REGION Network 178: %DB59.DBW2
   RUNG wire#powerrail
      I_Contact( "Rec_Todas" )
      I_Contact( "ResumAla_Grave" )
      { S7_GenerateENO := "TRUE" } Move(in := 0, out1 => %DB59.DBW2)
   END_RUNG
   // the same network as SCL:
   IF NOT "Rec_Todas" AND NOT "ResumAla_Grave" THEN %DB59.DBW2 := 0; END_IF;
END_REGION

REGION Network 179: %DB59.DBD4
   RUNG wire#powerrail
      Contact( "Rec_Todas" )
      wire#w1
      { S7_GenerateENO := "TRUE" } Move(in := DW#16#FFFFFFFF, out1 => %DB59.DBD4)
   END_RUNG
   RUNG wire#powerrail
      Contact( "ResumAla_Grave" )
   END_RUNG wire#w1
   // the same network as SCL:
   IF "Rec_Todas" OR "ResumAla_Grave" THEN %DB59.DBD4 := DW#16#FFFFFFFF; END_IF;
END_REGION

REGION Network 180: %DB59.DBD4
   RUNG wire#powerrail
      I_Contact( "Rec_Todas" )
      I_Contact( "ResumAla_Grave" )
      { S7_GenerateENO := "TRUE" } Move(in := 0, out1 => %DB59.DBD4)
   END_RUNG
   // the same network as SCL:
   IF NOT "Rec_Todas" AND NOT "ResumAla_Grave" THEN %DB59.DBD4 := 0; END_IF;
END_REGION

REGION Network 181: %DB59.DBD8
   RUNG wire#powerrail
      Contact( "Rec_Todas" )
      wire#w1
      { S7_GenerateENO := "TRUE" } Move(in := DW#16#FFFFFFFF, out1 => %DB59.DBD8)
   END_RUNG
   RUNG wire#powerrail
      Contact( "ResumAla_Grave" )
   END_RUNG wire#w1
   // the same network as SCL:
   IF "Rec_Todas" OR "ResumAla_Grave" THEN %DB59.DBD8 := DW#16#FFFFFFFF; END_IF;
END_REGION

REGION Network 182: %DB59.DBD8
   RUNG wire#powerrail
      I_Contact( "Rec_Todas" )
      I_Contact( "ResumAla_Grave" )
      { S7_GenerateENO := "TRUE" } Move(in := 0, out1 => %DB59.DBD8)
   END_RUNG
   // the same network as SCL:
   IF NOT "Rec_Todas" AND NOT "ResumAla_Grave" THEN %DB59.DBD8 := 0; END_IF;
END_REGION

REGION Network 183: %DB59.DBD12
   RUNG wire#powerrail
      Contact( "Rec_Todas" )
      wire#w1
      { S7_GenerateENO := "TRUE" } Move(in := DW#16#FFFFFFFF, out1 => %DB59.DBD12)
   END_RUNG
   RUNG wire#powerrail
      Contact( "ResumAla_Grave" )
   END_RUNG wire#w1
   // the same network as SCL:
   IF "Rec_Todas" OR "ResumAla_Grave" THEN %DB59.DBD12 := DW#16#FFFFFFFF; END_IF;
END_REGION

REGION Network 184: %DB59.DBD12
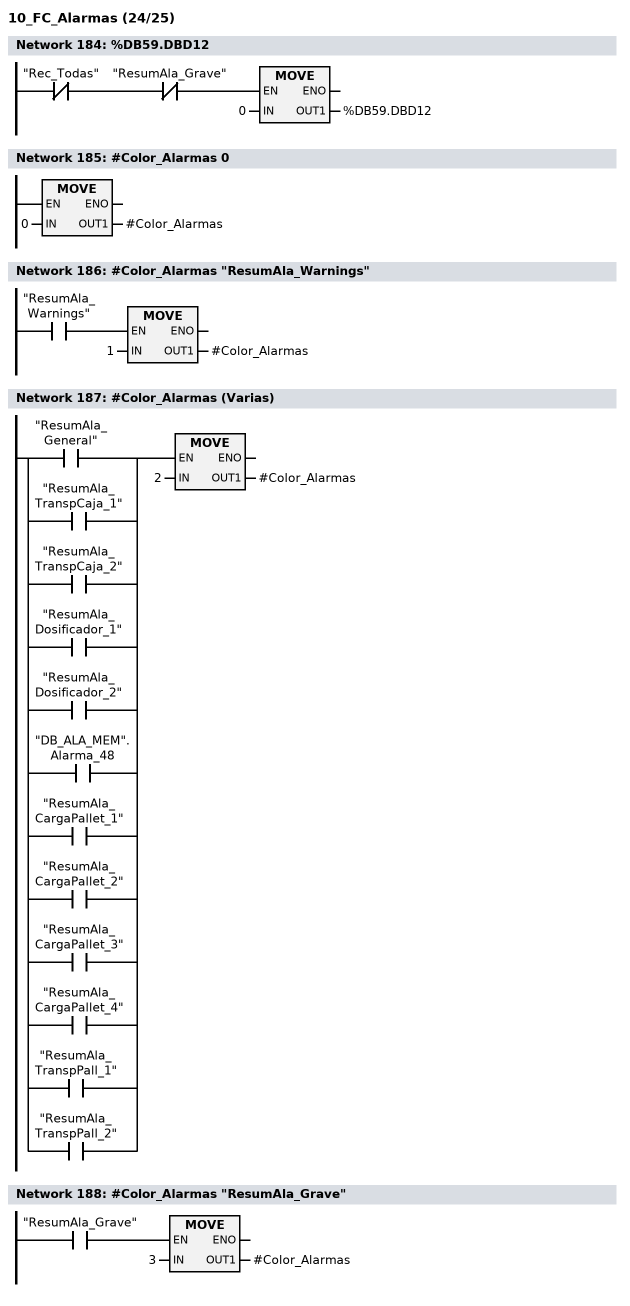
   RUNG wire#powerrail
      I_Contact( "Rec_Todas" )
      I_Contact( "ResumAla_Grave" )
      { S7_GenerateENO := "TRUE" } Move(in := 0, out1 => %DB59.DBD12)
   END_RUNG
   // the same network as SCL:
   IF NOT "Rec_Todas" AND NOT "ResumAla_Grave" THEN %DB59.DBD12 := 0; END_IF;
END_REGION

REGION Network 185: #Color_Alarmas 0
   RUNG wire#powerrail
      { S7_GenerateENO := "TRUE" } Move(in := 0, out1 => #Color_Alarmas)
   END_RUNG
   // the same network as SCL:
   #Color_Alarmas := 0;
END_REGION

REGION Network 186: #Color_Alarmas "ResumAla_Warnings"
   RUNG wire#powerrail
      Contact( "ResumAla_Warnings" )
      { S7_GenerateENO := "TRUE" } Move(in := 1, out1 => #Color_Alarmas)
   END_RUNG
   // the same network as SCL:
   IF "ResumAla_Warnings" THEN #Color_Alarmas := 1; END_IF;
END_REGION

REGION Network 187: #Color_Alarmas (Varias)
   RUNG wire#powerrail
      Contact( "ResumAla_General" )
      wire#w1
      { S7_GenerateENO := "TRUE" } Move(in := 2, out1 => #Color_Alarmas)
   END_RUNG
   RUNG wire#powerrail
      Contact( "ResumAla_TranspCaja_1" )
   END_RUNG wire#w1
   RUNG wire#powerrail
      Contact( "ResumAla_TranspCaja_2" )
   END_RUNG wire#w1
   RUNG wire#powerrail
      Contact( "ResumAla_Dosificador_1" )
   END_RUNG wire#w1
   RUNG wire#powerrail
      Contact( "ResumAla_Dosificador_2" )
   END_RUNG wire#w1
   RUNG wire#powerrail
      Contact( "DB_ALA_MEM".Alarma_48 )
   END_RUNG wire#w1
   RUNG wire#powerrail
      Contact( "ResumAla_CargaPallet_1" )
   END_RUNG wire#w1
   RUNG wire#powerrail
      Contact( "ResumAla_CargaPallet_2" )
   END_RUNG wire#w1
   RUNG wire#powerrail
      Contact( "ResumAla_CargaPallet_3" )
   END_RUNG wire#w1
   RUNG wire#powerrail
      Contact( "ResumAla_CargaPallet_4" )
   END_RUNG wire#w1
   RUNG wire#powerrail
      Contact( "ResumAla_TranspPall_1" )
   END_RUNG wire#w1
   RUNG wire#powerrail
      Contact( "ResumAla_TranspPall_2" )
   END_RUNG wire#w1
   // the same network as SCL:
   IF "ResumAla_General" OR "ResumAla_TranspCaja_1" OR "ResumAla_TranspCaja_2" OR "ResumAla_Dosificador_1" OR "ResumAla_Dosificador_2" OR "DB_ALA_MEM".Alarma_48 OR "ResumAla_CargaPallet_1" OR "ResumAla_CargaPallet_2" OR "ResumAla_CargaPallet_3" OR "ResumAla_CargaPallet_4" OR "ResumAla_TranspPall_1" OR "ResumAla_TranspPall_2" THEN
       #Color_Alarmas := 2;
   END_IF;
END_REGION

REGION Network 188: #Color_Alarmas "ResumAla_Grave"
   RUNG wire#powerrail
      Contact( "ResumAla_Grave" )
      { S7_GenerateENO := "TRUE" } Move(in := 3, out1 => #Color_Alarmas)
   END_RUNG
   // the same network as SCL:
   IF "ResumAla_Grave" THEN #Color_Alarmas := 3; END_IF;
END_REGION

REGION Network 189: "Color_Alarmas"
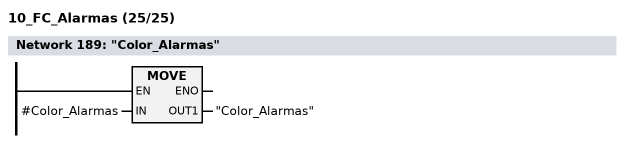
   RUNG wire#powerrail
      { S7_GenerateENO := "TRUE" } Move(in := #Color_Alarmas, out1 => "Color_Alarmas")
   END_RUNG
   // the same network as SCL:
   "Color_Alarmas" := #Color_Alarmas;
END_REGION
END_FUNCTION

// folder: Estandar

FUNCTION_BLOCK "FB_VAR_MOT"   // FB2, LAD
{ S7_Optimized_Access := 'FALSE' }
VERSION : 0.1
   VAR_TEMP   // added for the SCL form of the ladder/FBD networks
      _w1 : Bool;
      _w2 : Bool;
      _w3 : Bool;
   END_VAR
BEGIN

REGION Network 1: #Aux
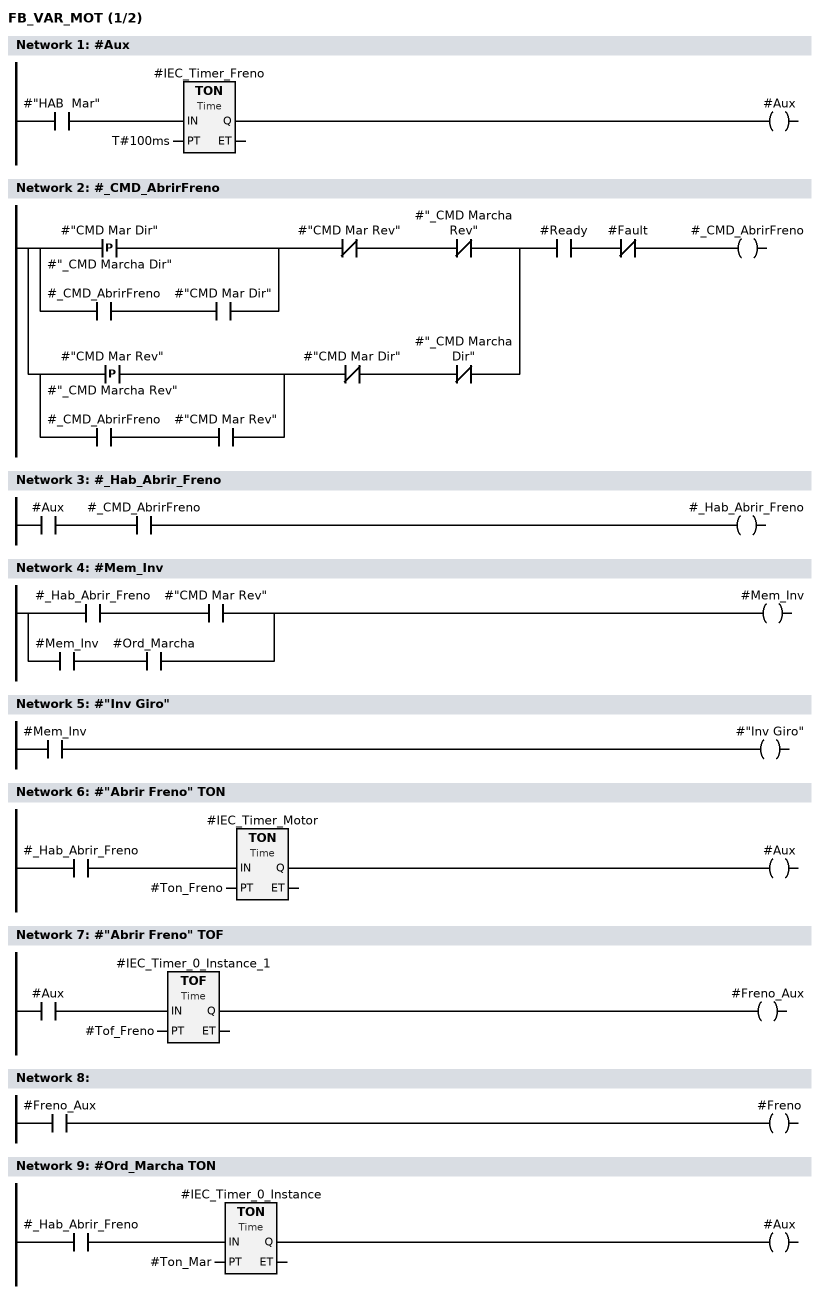
   #IEC_Timer_Freno.TON(in := #"HAB  Mar", pt := T#100ms);
   #Aux := #IEC_Timer_Freno.q;
END_REGION

REGION Network 2: #_CMD_AbrirFreno
   RUNG wire#powerrail
      P_Contact(operand := #"CMD Mar Dir", bit := #"_CMD Marcha Dir")
      wire#w1
      I_Contact( #"CMD Mar Rev" )
      I_Contact( #"_CMD Marcha Rev" )
      wire#w2
      Contact( #Ready )
      I_Contact( #Fault )
      Coil( #_CMD_AbrirFreno )
   END_RUNG
   RUNG wire#powerrail
      Contact( #_CMD_AbrirFreno )
      Contact( #"CMD Mar Dir" )
   END_RUNG wire#w1
   RUNG wire#powerrail
      P_Contact(operand := #"CMD Mar Rev", bit := #"_CMD Marcha Rev")
      wire#w3
      I_Contact( #"CMD Mar Dir" )
      I_Contact( #"_CMD Marcha Dir" )
   END_RUNG wire#w2
   RUNG wire#powerrail
      Contact( #_CMD_AbrirFreno )
      Contact( #"CMD Mar Rev" )
   END_RUNG wire#w3
   // the same network as SCL:
   #_w1 := #"CMD Mar Dir" AND NOT #"_CMD Marcha Dir";   // rising edge of #"CMD Mar Dir"
   #"_CMD Marcha Dir" := #"CMD Mar Dir";
   #_w3 := (#_w1 OR (#_CMD_AbrirFreno AND #"CMD Mar Dir")) AND NOT #"CMD Mar Rev" AND NOT #"_CMD Marcha Rev";
   #_w2 := #"CMD Mar Rev" AND NOT #"_CMD Marcha Rev";   // rising edge of #"CMD Mar Rev"
   #"_CMD Marcha Rev" := #"CMD Mar Rev";
   #_CMD_AbrirFreno := (#_w3 OR ((#_w2 OR (#_CMD_AbrirFreno AND #"CMD Mar Rev")) AND NOT #"CMD Mar Dir" AND NOT #"_CMD Marcha Dir")) AND #Ready AND NOT #Fault;
END_REGION

REGION Network 3: #_Hab_Abrir_Freno
   RUNG wire#powerrail
      Contact( #Aux )
      Contact( #_CMD_AbrirFreno )
      Coil( #_Hab_Abrir_Freno )
   END_RUNG
   // the same network as SCL:
   #_Hab_Abrir_Freno := #Aux AND #_CMD_AbrirFreno;
END_REGION

REGION Network 4: #Mem_Inv
   RUNG wire#powerrail
      Contact( #_Hab_Abrir_Freno )
      Contact( #"CMD Mar Rev" )
      wire#w1
      Coil( #Mem_Inv )
   END_RUNG
   RUNG wire#powerrail
      Contact( #Mem_Inv )
      Contact( #Ord_Marcha )
   END_RUNG wire#w1
   // the same network as SCL:
   #Mem_Inv := (#_Hab_Abrir_Freno AND #"CMD Mar Rev") OR (#Mem_Inv AND #Ord_Marcha);
END_REGION

REGION Network 5: #"Inv Giro"
   RUNG wire#powerrail
      Contact( #Mem_Inv )
      Coil( #"Inv Giro" )
   END_RUNG
   // the same network as SCL:
   #"Inv Giro" := #Mem_Inv;
END_REGION

REGION Network 6: #"Abrir Freno" TON
   #IEC_Timer_Motor.TON(in := #_Hab_Abrir_Freno, pt := #Ton_Freno);
   #Aux := #IEC_Timer_Motor.q;
END_REGION

REGION Network 7: #"Abrir Freno" TOF
   #IEC_Timer_0_Instance_1.TOF(in := #Aux, pt := #Tof_Freno);
   #Freno_Aux := #IEC_Timer_0_Instance_1.q;
END_REGION

REGION Network 8
   RUNG wire#powerrail
      Contact( #Freno_Aux )
      Coil( #Freno )
   END_RUNG
   // the same network as SCL:
   #Freno := #Freno_Aux;
END_REGION

REGION Network 9: #Ord_Marcha TON
   #IEC_Timer_0_Instance.TON(in := #_Hab_Abrir_Freno, pt := #Ton_Mar);
   #Aux := #IEC_Timer_0_Instance.q;
END_REGION

REGION Network 10: #Ord_Marcha TOF
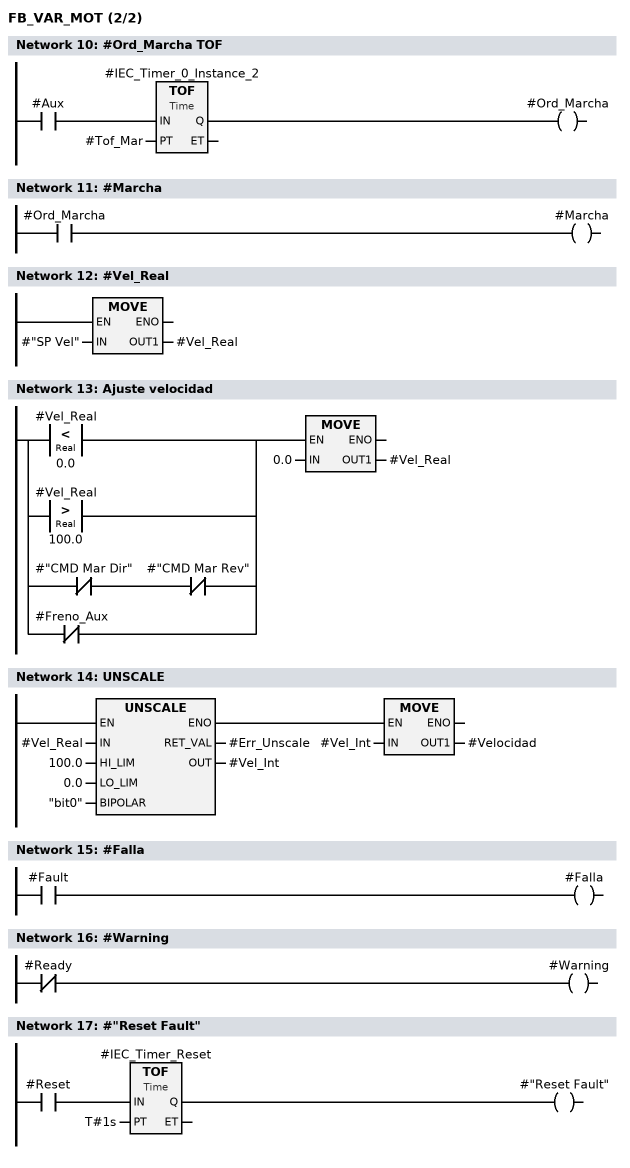
   #IEC_Timer_0_Instance_2.TOF(in := #Aux, pt := #Tof_Mar);
   #Ord_Marcha := #IEC_Timer_0_Instance_2.q;
END_REGION

REGION Network 11: #Marcha
   RUNG wire#powerrail
      Contact( #Ord_Marcha )
      Coil( #Marcha )
   END_RUNG
   // the same network as SCL:
   #Marcha := #Ord_Marcha;
END_REGION

REGION Network 12: #Vel_Real
   RUNG wire#powerrail
      { S7_GenerateENO := "TRUE" } Move(in := #"SP Vel", out1 => #Vel_Real)
   END_RUNG
   // the same network as SCL:
   #Vel_Real := #"SP Vel";
END_REGION

REGION Network 13: Ajuste velocidad
   RUNG wire#powerrail
      { S7_Templates := "SrcType := Real" } LT_Contact(in1 := #Vel_Real, in2 := 0.0)
      wire#w1
      { S7_GenerateENO := "TRUE" } Move(in := 0.0, out1 => #Vel_Real)
   END_RUNG
   RUNG wire#powerrail
      { S7_Templates := "SrcType := Real" } GT_Contact(in1 := #Vel_Real, in2 := 100.0)
   END_RUNG wire#w1
   RUNG wire#powerrail
      I_Contact( #"CMD Mar Dir" )
      I_Contact( #"CMD Mar Rev" )
   END_RUNG wire#w1
   RUNG wire#powerrail
      I_Contact( #Freno_Aux )
   END_RUNG wire#w1
   // the same network as SCL:
   IF (#Vel_Real < 0.0) OR (#Vel_Real > 100.0) OR (NOT #"CMD Mar Dir" AND NOT #"CMD Mar Rev") OR NOT #Freno_Aux THEN
       #Vel_Real := 0.0;
   END_IF;
END_REGION

REGION Network 14: UNSCALE
   // ENO of a box is taken as its EN; it also drops when the box reports an error
   #Err_Unscale := UNSCALE(in := #Vel_Real, hi_lim := 100.0, lo_lim := 0.0, bipolar := "bit0", out => #Vel_Int);
   #Velocidad := #Vel_Int;
END_REGION

REGION Network 15: #Falla
   RUNG wire#powerrail
      Contact( #Fault )
      Coil( #Falla )
   END_RUNG
   // the same network as SCL:
   #Falla := #Fault;
END_REGION

REGION Network 16: #Warning
   RUNG wire#powerrail
      I_Contact( #Ready )
      Coil( #Warning )
   END_RUNG
   // the same network as SCL:
   #Warning := NOT #Ready;
END_REGION

REGION Network 17: #"Reset Fault"
   #IEC_Timer_Reset.TOF(in := #Reset, pt := T#1s);
   #"Reset Fault" := #IEC_Timer_Reset.q;
END_REGION
END_FUNCTION_BLOCK

FUNCTION_BLOCK "FB_CTR_VAL"   // FB3, LAD
{ S7_Optimized_Access := 'FALSE' }
VERSION : 0.1
BEGIN

REGION Network 1: #_CMD
   // Si no está habilitado mantiene el estado anterior
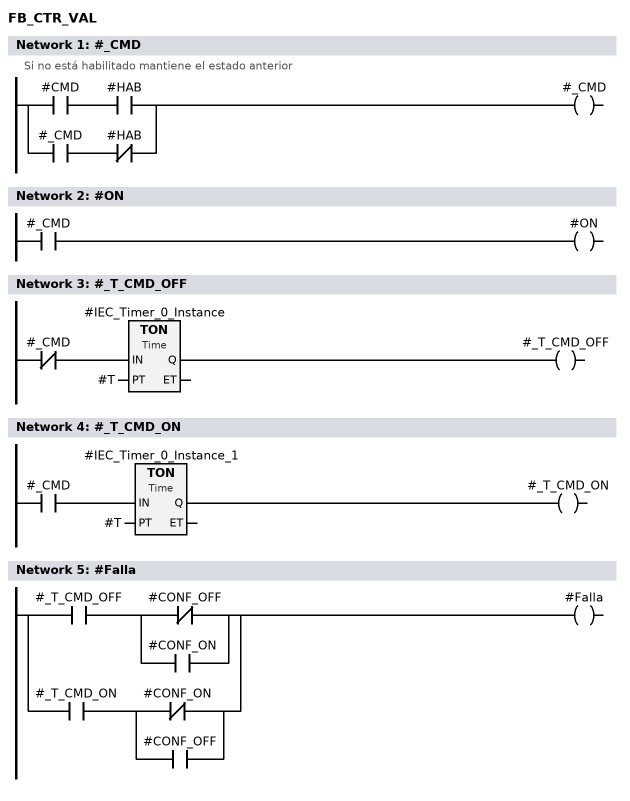
   RUNG wire#powerrail
      Contact( #CMD )
      Contact( #HAB )
      wire#w1
      Coil( #_CMD )
   END_RUNG
   RUNG wire#powerrail
      Contact( #_CMD )
      I_Contact( #HAB )
   END_RUNG wire#w1
   // the same network as SCL:
   #_CMD := (#CMD AND #HAB) OR (#_CMD AND NOT #HAB);
END_REGION

REGION Network 2: #ON
   RUNG wire#powerrail
      Contact( #_CMD )
      Coil( #ON )
   END_RUNG
   // the same network as SCL:
   #ON := #_CMD;
END_REGION

REGION Network 3: #_T_CMD_OFF
   #IEC_Timer_0_Instance.TON(in := NOT #_CMD, pt := #T);
   #_T_CMD_OFF := #IEC_Timer_0_Instance.q;
END_REGION

REGION Network 4: #_T_CMD_ON
   #IEC_Timer_0_Instance_1.TON(in := #_CMD, pt := #T);
   #_T_CMD_ON := #IEC_Timer_0_Instance_1.q;
END_REGION

REGION Network 5: #Falla
   RUNG wire#powerrail
      Contact( #_T_CMD_OFF )
      wire#w1
      I_Contact( #CONF_OFF )
      wire#w2
      Coil( #Falla )
   END_RUNG
   RUNG wire#w1
      Contact( #CONF_ON )
   END_RUNG wire#w2
   RUNG wire#powerrail
      Contact( #_T_CMD_ON )
      wire#w3
      I_Contact( #CONF_ON )
   END_RUNG wire#w2
   RUNG wire#w3
      Contact( #CONF_OFF )
   END_RUNG wire#w2
   // the same network as SCL:
   #Falla := (#_T_CMD_OFF AND (NOT #CONF_OFF OR #CONF_ON)) OR (#_T_CMD_ON AND (NOT #CONF_ON OR #CONF_OFF));
END_REGION
END_FUNCTION_BLOCK

FUNCTION_BLOCK "FB_CTR_MOT_FRD"   // FB4, LAD
{ S7_Optimized_Access := 'FALSE' }
VERSION : 0.1
   VAR_TEMP   // added for the SCL form of the ladder/FBD networks
      _w1 : Bool;
      _w2 : Bool;
      _w3 : Bool;
   END_VAR
BEGIN

REGION Network 1: #_REQ_Marcha
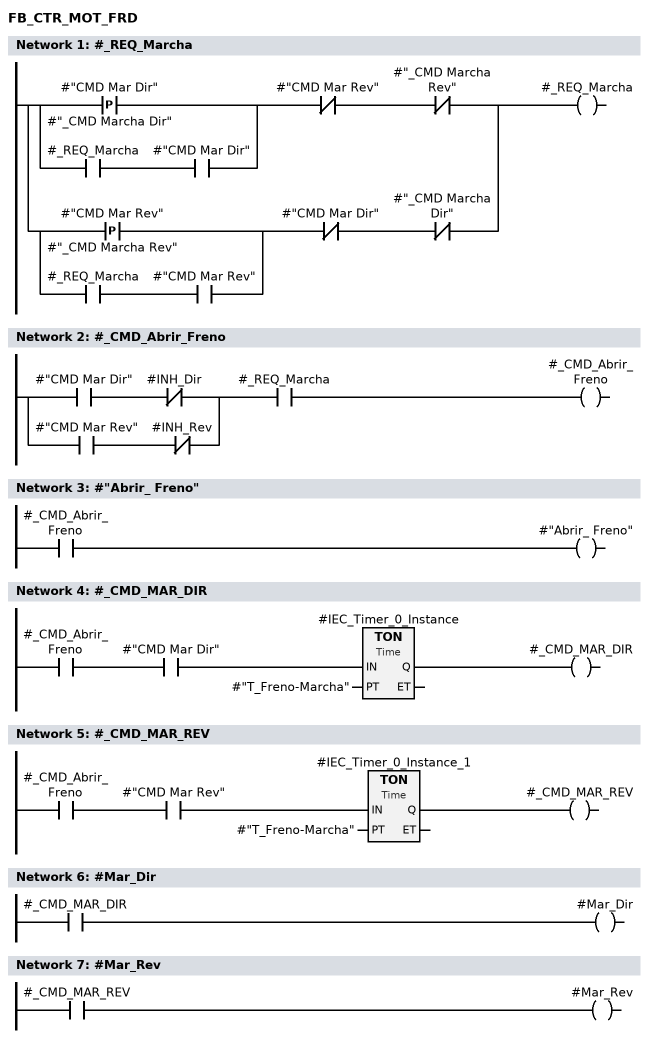
   RUNG wire#powerrail
      P_Contact(operand := #"CMD Mar Dir", bit := #"_CMD Marcha Dir")
      wire#w1
      I_Contact( #"CMD Mar Rev" )
      I_Contact( #"_CMD Marcha Rev" )
      wire#w2
      Coil( #_REQ_Marcha )
   END_RUNG
   RUNG wire#powerrail
      Contact( #_REQ_Marcha )
      Contact( #"CMD Mar Dir" )
   END_RUNG wire#w1
   RUNG wire#powerrail
      P_Contact(operand := #"CMD Mar Rev", bit := #"_CMD Marcha Rev")
      wire#w3
      I_Contact( #"CMD Mar Dir" )
      I_Contact( #"_CMD Marcha Dir" )
   END_RUNG wire#w2
   RUNG wire#powerrail
      Contact( #_REQ_Marcha )
      Contact( #"CMD Mar Rev" )
   END_RUNG wire#w3
   // the same network as SCL:
   #_w1 := #"CMD Mar Dir" AND NOT #"_CMD Marcha Dir";   // rising edge of #"CMD Mar Dir"
   #"_CMD Marcha Dir" := #"CMD Mar Dir";
   #_w3 := (#_w1 OR (#_REQ_Marcha AND #"CMD Mar Dir")) AND NOT #"CMD Mar Rev" AND NOT #"_CMD Marcha Rev";
   #_w2 := #"CMD Mar Rev" AND NOT #"_CMD Marcha Rev";   // rising edge of #"CMD Mar Rev"
   #"_CMD Marcha Rev" := #"CMD Mar Rev";
   #_REQ_Marcha := #_w3 OR ((#_w2 OR (#_REQ_Marcha AND #"CMD Mar Rev")) AND NOT #"CMD Mar Dir" AND NOT #"_CMD Marcha Dir");
END_REGION

REGION Network 2: #_CMD_Abrir_Freno
   RUNG wire#powerrail
      Contact( #"CMD Mar Dir" )
      I_Contact( #INH_Dir )
      wire#w1
      Contact( #_REQ_Marcha )
      Coil( #_CMD_Abrir_Freno )
   END_RUNG
   RUNG wire#powerrail
      Contact( #"CMD Mar Rev" )
      I_Contact( #INH_Rev )
   END_RUNG wire#w1
   // the same network as SCL:
   #_CMD_Abrir_Freno := ((#"CMD Mar Dir" AND NOT #INH_Dir) OR (#"CMD Mar Rev" AND NOT #INH_Rev)) AND #_REQ_Marcha;
END_REGION

REGION Network 3: #"Abrir_ Freno"
   RUNG wire#powerrail
      Contact( #_CMD_Abrir_Freno )
      Coil( #"Abrir_ Freno" )
   END_RUNG
   // the same network as SCL:
   #"Abrir_ Freno" := #_CMD_Abrir_Freno;
END_REGION

REGION Network 4: #_CMD_MAR_DIR
   #IEC_Timer_0_Instance.TON(in := #_CMD_Abrir_Freno AND #"CMD Mar Dir", pt := #"T_Freno-Marcha");
   #_CMD_MAR_DIR := #IEC_Timer_0_Instance.q;
END_REGION

REGION Network 5: #_CMD_MAR_REV
   #IEC_Timer_0_Instance_1.TON(in := #_CMD_Abrir_Freno AND #"CMD Mar Rev", pt := #"T_Freno-Marcha");
   #_CMD_MAR_REV := #IEC_Timer_0_Instance_1.q;
END_REGION

REGION Network 6: #Mar_Dir
   RUNG wire#powerrail
      Contact( #_CMD_MAR_DIR )
      Coil( #Mar_Dir )
   END_RUNG
   // the same network as SCL:
   #Mar_Dir := #_CMD_MAR_DIR;
END_REGION

REGION Network 7: #Mar_Rev
   RUNG wire#powerrail
      Contact( #_CMD_MAR_REV )
      Coil( #Mar_Rev )
   END_RUNG
   // the same network as SCL:
   #Mar_Rev := #_CMD_MAR_REV;
END_REGION
END_FUNCTION_BLOCK

// folder: Grupos

FUNCTION "3_FC_Transp_Cajas" : Void   // FC7, LAD
{ S7_Optimized_Access := 'FALSE' }
VERSION : 0.1
BEGIN

REGION Network 1: Resets "HMI".Pls_MarMan_R...
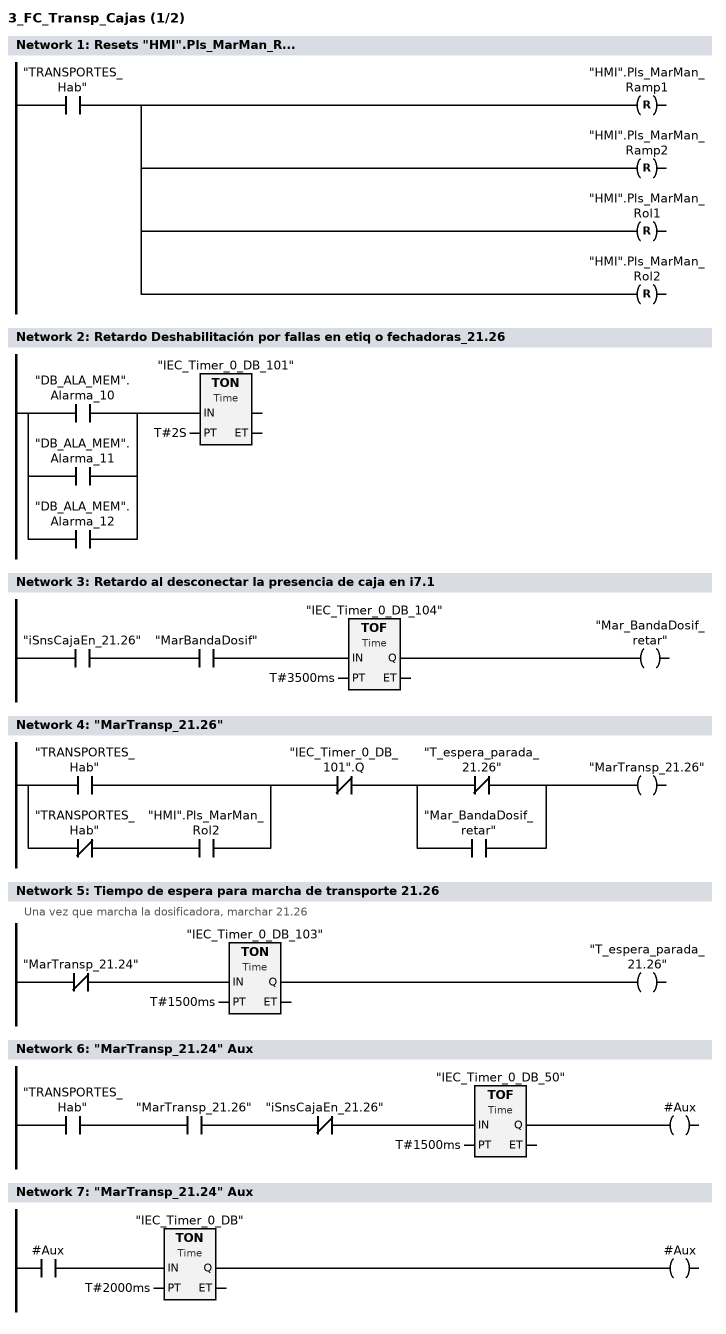
   RUNG wire#powerrail
      Contact( "TRANSPORTES_Hab" )
      wire#w1
      R_Coil( "HMI".Pls_MarMan_Ramp1 )
   END_RUNG
   RUNG wire#w1
      R_Coil( "HMI".Pls_MarMan_Ramp2 )
   END_RUNG
   RUNG wire#w1
      R_Coil( "HMI".Pls_MarMan_Rol1 )
   END_RUNG
   RUNG wire#w1
      R_Coil( "HMI".Pls_MarMan_Rol2 )
   END_RUNG
   // the same network as SCL:
   IF "TRANSPORTES_Hab" THEN
       "HMI".Pls_MarMan_Ramp1 := FALSE;
       "HMI".Pls_MarMan_Ramp2 := FALSE;
       "HMI".Pls_MarMan_Rol1 := FALSE;
       "HMI".Pls_MarMan_Rol2 := FALSE;
   END_IF;
END_REGION

REGION Network 2: Retardo Deshabilitación por fallas en etiq o fechadoras_21.26
   "IEC_Timer_0_DB_101".TON(IN := "DB_ALA_MEM".Alarma_10 OR "DB_ALA_MEM".Alarma_11 OR "DB_ALA_MEM".Alarma_12,
                           PT := T#2S);
END_REGION

REGION Network 3: Retardo al desconectar la presencia de caja en i7.1
   "IEC_Timer_0_DB_104".TOF(IN := "iSnsCajaEn_21.26" AND "MarBandaDosif", PT := T#3500ms);
   "Mar_BandaDosif_retar" := "IEC_Timer_0_DB_104".Q;
END_REGION

REGION Network 4: "MarTransp_21.26"
   RUNG wire#powerrail
      Contact( "TRANSPORTES_Hab" )
      wire#w1
      I_Contact( "IEC_Timer_0_DB_101".Q )
      wire#w2
      I_Contact( "T_espera_parada_21.26" )
      wire#w3
      Coil( "MarTransp_21.26" )
   END_RUNG
   RUNG wire#powerrail
      I_Contact( "TRANSPORTES_Hab" )
      Contact( "HMI".Pls_MarMan_Rol2 )
   END_RUNG wire#w1
   RUNG wire#w2
      Contact( "Mar_BandaDosif_retar" )
   END_RUNG wire#w3
   // the same network as SCL:
   "MarTransp_21.26" := ("TRANSPORTES_Hab" OR (NOT "TRANSPORTES_Hab" AND "HMI".Pls_MarMan_Rol2)) AND NOT "IEC_Timer_0_DB_101".Q AND (NOT "T_espera_parada_21.26" OR "Mar_BandaDosif_retar");
END_REGION

REGION Network 5: Tiempo de espera para marcha de transporte 21.26
   // Una vez que marcha la dosificadora, marchar 21.26
   "IEC_Timer_0_DB_103".TON(IN := NOT "MarTransp_21.24", PT := T#1500ms);
   "T_espera_parada_21.26" := "IEC_Timer_0_DB_103".Q;
END_REGION

REGION Network 6: "MarTransp_21.24" Aux
   "IEC_Timer_0_DB_50".TOF(IN := "TRANSPORTES_Hab" AND "MarTransp_21.26" AND NOT "iSnsCajaEn_21.26",
                           PT := T#1500ms);
   #Aux := "IEC_Timer_0_DB_50".Q;
END_REGION

REGION Network 7: "MarTransp_21.24" Aux
   "IEC_Timer_0_DB".TON(IN := #Aux, PT := T#2000ms);
   #Aux := "IEC_Timer_0_DB".Q;
END_REGION

REGION Network 8: "MarTransp_21.24"
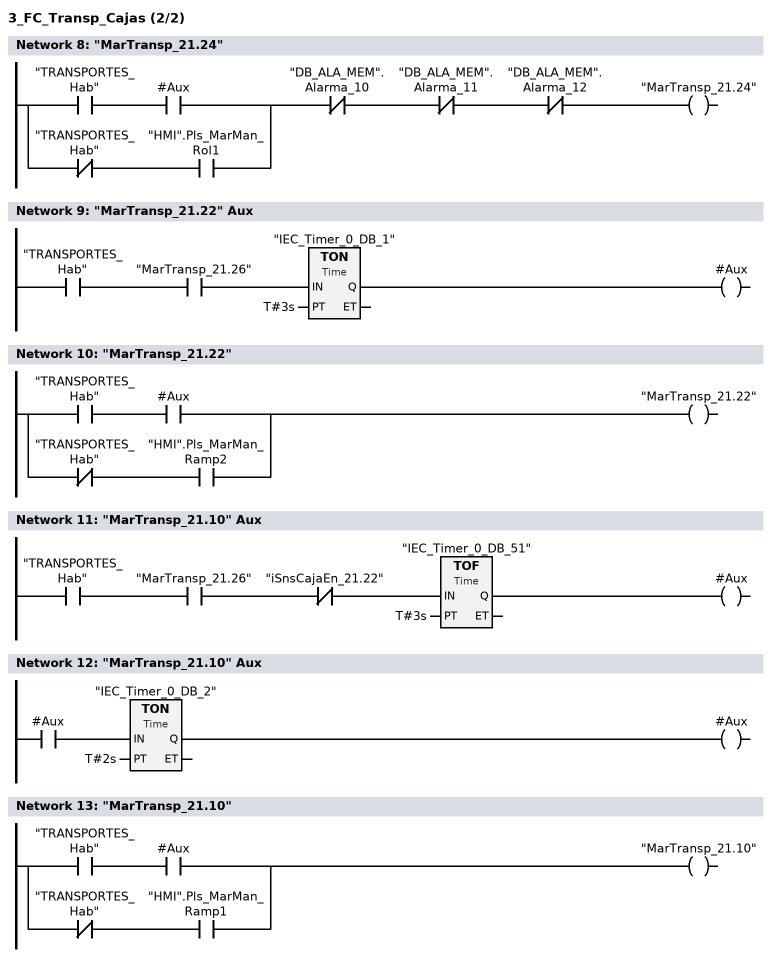
   RUNG wire#powerrail
      Contact( "TRANSPORTES_Hab" )
      Contact( #Aux )
      wire#w1
      I_Contact( "DB_ALA_MEM".Alarma_10 )
      I_Contact( "DB_ALA_MEM".Alarma_11 )
      I_Contact( "DB_ALA_MEM".Alarma_12 )
      Coil( "MarTransp_21.24" )
   END_RUNG
   RUNG wire#powerrail
      I_Contact( "TRANSPORTES_Hab" )
      Contact( "HMI".Pls_MarMan_Rol1 )
   END_RUNG wire#w1
   // the same network as SCL:
   "MarTransp_21.24" := (("TRANSPORTES_Hab" AND #Aux) OR (NOT "TRANSPORTES_Hab" AND "HMI".Pls_MarMan_Rol1)) AND NOT "DB_ALA_MEM".Alarma_10 AND NOT "DB_ALA_MEM".Alarma_11 AND NOT "DB_ALA_MEM".Alarma_12;
END_REGION

REGION Network 9: "MarTransp_21.22" Aux
   "IEC_Timer_0_DB_1".TON(IN := "TRANSPORTES_Hab" AND "MarTransp_21.26", PT := T#3s);
   #Aux := "IEC_Timer_0_DB_1".Q;
END_REGION

REGION Network 10: "MarTransp_21.22"
   RUNG wire#powerrail
      Contact( "TRANSPORTES_Hab" )
      Contact( #Aux )
      wire#w1
      Coil( "MarTransp_21.22" )
   END_RUNG
   RUNG wire#powerrail
      I_Contact( "TRANSPORTES_Hab" )
      Contact( "HMI".Pls_MarMan_Ramp2 )
   END_RUNG wire#w1
   // the same network as SCL:
   "MarTransp_21.22" := ("TRANSPORTES_Hab" AND #Aux) OR (NOT "TRANSPORTES_Hab" AND "HMI".Pls_MarMan_Ramp2);
END_REGION

REGION Network 11: "MarTransp_21.10" Aux
   "IEC_Timer_0_DB_51".TOF(IN := "TRANSPORTES_Hab" AND "MarTransp_21.26" AND NOT "iSnsCajaEn_21.22", PT := T#3s);
   #Aux := "IEC_Timer_0_DB_51".Q;
END_REGION

REGION Network 12: "MarTransp_21.10" Aux
   "IEC_Timer_0_DB_2".TON(IN := #Aux, PT := T#2s);
   #Aux := "IEC_Timer_0_DB_2".Q;
END_REGION

REGION Network 13: "MarTransp_21.10"
   RUNG wire#powerrail
      Contact( "TRANSPORTES_Hab" )
      Contact( #Aux )
      wire#w1
      Coil( "MarTransp_21.10" )
   END_RUNG
   RUNG wire#powerrail
      I_Contact( "TRANSPORTES_Hab" )
      Contact( "HMI".Pls_MarMan_Ramp1 )
   END_RUNG wire#w1
   // the same network as SCL:
   "MarTransp_21.10" := ("TRANSPORTES_Hab" AND #Aux) OR (NOT "TRANSPORTES_Hab" AND "HMI".Pls_MarMan_Ramp1);
END_REGION
END_FUNCTION

FUNCTION "2_FC_General" : Void   // FC8, LAD
{ S7_Optimized_Access := 'FALSE' }
VERSION : 0.1
   VAR_TEMP   // added for the SCL form of the ladder/FBD networks
      _w1 : Bool;
   END_VAR
BEGIN

REGION Network 1: "AUTO/MAN"
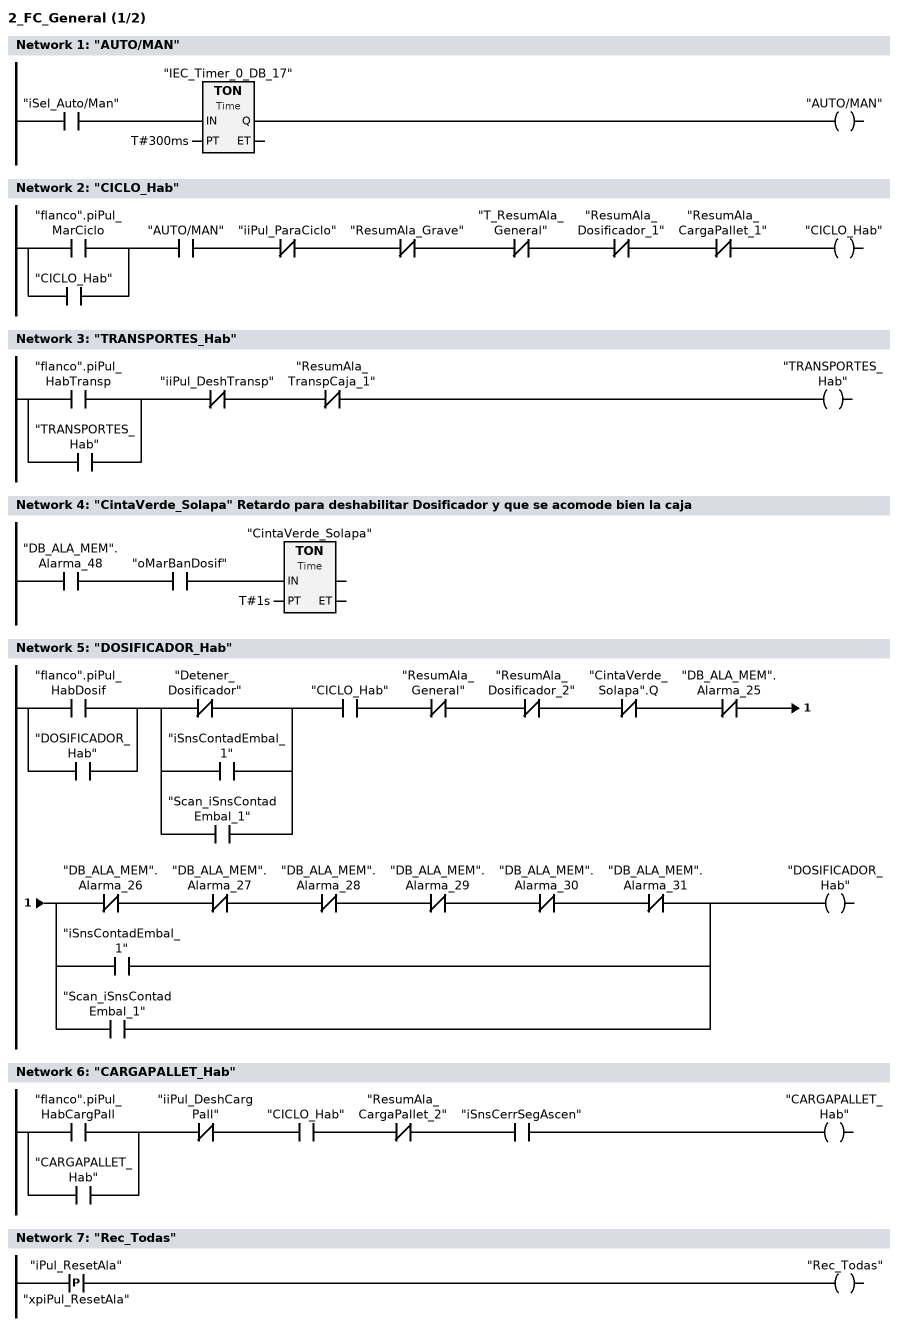
   "IEC_Timer_0_DB_17".TON(in := "iSel_Auto/Man", pt := T#300ms);
   "AUTO/MAN" := "IEC_Timer_0_DB_17".q;
END_REGION

REGION Network 2: "CICLO_Hab"
   RUNG wire#powerrail
      Contact( "flanco".piPul_MarCiclo )
      wire#w1
      Contact( "AUTO/MAN" )
      I_Contact( "iiPul_ParaCiclo" )
      I_Contact( "ResumAla_Grave" )
      I_Contact( "T_ResumAla_General" )
      I_Contact( "ResumAla_Dosificador_1" )
      I_Contact( "ResumAla_CargaPallet_1" )
      Coil( "CICLO_Hab" )
   END_RUNG
   RUNG wire#powerrail
      Contact( "CICLO_Hab" )
   END_RUNG wire#w1
   // the same network as SCL:
   "CICLO_Hab" := ("flanco".piPul_MarCiclo OR "CICLO_Hab") AND "AUTO/MAN" AND NOT "iiPul_ParaCiclo" AND NOT "ResumAla_Grave" AND NOT "T_ResumAla_General" AND NOT "ResumAla_Dosificador_1" AND NOT "ResumAla_CargaPallet_1";
END_REGION

REGION Network 3: "TRANSPORTES_Hab"
   RUNG wire#powerrail
      Contact( "flanco".piPul_HabTransp )
      wire#w1
      I_Contact( "iiPul_DeshTransp" )
      I_Contact( "ResumAla_TranspCaja_1" )
      Coil( "TRANSPORTES_Hab" )
   END_RUNG
   RUNG wire#powerrail
      Contact( "TRANSPORTES_Hab" )
   END_RUNG wire#w1
   // the same network as SCL:
   "TRANSPORTES_Hab" := ("flanco".piPul_HabTransp OR "TRANSPORTES_Hab") AND NOT "iiPul_DeshTransp" AND NOT "ResumAla_TranspCaja_1";
END_REGION

REGION Network 4: "CintaVerde_Solapa" Retardo para deshabilitar Dosificador y que se acomode bien la caja
   "CintaVerde_Solapa".TON(IN := "DB_ALA_MEM".Alarma_48 AND "oMarBanDosif", PT := T#1s);
END_REGION

REGION Network 5: "DOSIFICADOR_Hab"
   RUNG wire#powerrail
      Contact( "flanco".piPul_HabDosif )
      wire#w1
      I_Contact( "Detener_Dosificador" )
      wire#w2
      Contact( "CICLO_Hab" )
      I_Contact( "ResumAla_General" )
      I_Contact( "ResumAla_Dosificador_2" )
      I_Contact( "CintaVerde_Solapa".Q )
      I_Contact( "DB_ALA_MEM".Alarma_25 )
      wire#w3
      I_Contact( "DB_ALA_MEM".Alarma_26 )
      I_Contact( "DB_ALA_MEM".Alarma_27 )
      I_Contact( "DB_ALA_MEM".Alarma_28 )
      I_Contact( "DB_ALA_MEM".Alarma_29 )
      I_Contact( "DB_ALA_MEM".Alarma_30 )
      I_Contact( "DB_ALA_MEM".Alarma_31 )
      wire#w4
      Coil( "DOSIFICADOR_Hab" )
   END_RUNG
   RUNG wire#powerrail
      Contact( "DOSIFICADOR_Hab" )
   END_RUNG wire#w1
   RUNG wire#w1
      Contact( "iSnsContadEmbal_1" )
   END_RUNG wire#w2
   RUNG wire#w1
      Contact( "Scan_iSnsContadEmbal_1" )
   END_RUNG wire#w2
   RUNG wire#w3
      Contact( "iSnsContadEmbal_1" )
   END_RUNG wire#w4
   RUNG wire#w3
      Contact( "Scan_iSnsContadEmbal_1" )
   END_RUNG wire#w4
   // the same network as SCL:
   "DOSIFICADOR_Hab" := ("flanco".piPul_HabDosif OR "DOSIFICADOR_Hab") AND (NOT "Detener_Dosificador" OR "iSnsContadEmbal_1" OR "Scan_iSnsContadEmbal_1") AND "CICLO_Hab" AND NOT "ResumAla_General" AND NOT "ResumAla_Dosificador_2" AND NOT "CintaVerde_Solapa".Q AND NOT "DB_ALA_MEM".Alarma_25 AND ((NOT "DB_ALA_MEM".Alarma_26 AND NOT "DB_ALA_MEM".Alarma_27 AND NOT "DB_ALA_MEM".Alarma_28 AND NOT "DB_ALA_MEM".Alarma_29 AND NOT "DB_ALA_MEM".Alarma_30 AND NOT "DB_ALA_MEM".Alarma_31) OR "iSnsContadEmbal_1" OR "Scan_iSnsContadEmbal_1");
END_REGION

REGION Network 6: "CARGAPALLET_Hab"
   RUNG wire#powerrail
      Contact( "flanco".piPul_HabCargPall )
      wire#w1
      I_Contact( "iiPul_DeshCargPall" )
      Contact( "CICLO_Hab" )
      I_Contact( "ResumAla_CargaPallet_2" )
      Contact( "iSnsCerrSegAscen" )
      Coil( "CARGAPALLET_Hab" )
   END_RUNG
   RUNG wire#powerrail
      Contact( "CARGAPALLET_Hab" )
   END_RUNG wire#w1
   // the same network as SCL:
   "CARGAPALLET_Hab" := ("flanco".piPul_HabCargPall OR "CARGAPALLET_Hab") AND NOT "iiPul_DeshCargPall" AND "CICLO_Hab" AND NOT "ResumAla_CargaPallet_2" AND "iSnsCerrSegAscen";
END_REGION

REGION Network 7: "Rec_Todas"
   RUNG wire#powerrail
      P_Contact(operand := "iPul_ResetAla", bit := "xpiPul_ResetAla")
      Coil( "Rec_Todas" )
   END_RUNG
   // the same network as SCL:
   #_w1 := "iPul_ResetAla" AND NOT "xpiPul_ResetAla";   // rising edge of "iPul_ResetAla"
   "xpiPul_ResetAla" := "iPul_ResetAla";
   "Rec_Todas" := #_w1;
END_REGION

REGION Network 8: Imagen AUTO
